// TIA Portal project "Inteligenta_szklarnia" (V15.1) (continued)
REGION Network 5
   RUNG wire#powerrail
      "Rolety"(Czy_automatyczny := wire#w1, Czy_manualny := wire#w2)
   END_RUNG
   RUNG wire#powerrail
      Contact( "HMI".Aktywacja_trybu_automatycznego )
   END_RUNG wire#w1
   RUNG wire#powerrail
      Contact( "HMI".Aktywacja_trybu_manualnego )
   END_RUNG wire#w2
   // the same network as SCL:
   "Rolety"(Czy_automatyczny := "HMI".Aktywacja_trybu_automatycznego,
            Czy_manualny := "HMI".Aktywacja_trybu_manualnego);
END_REGION

REGION Network 6
   RUNG wire#powerrail
      "Zapis_parametrow_trybu_auto"()
   END_RUNG
   // the same network as SCL:
   "Zapis_parametrow_trybu_auto"();
END_REGION

REGION Network 7
   RUNG wire#powerrail
      P_Contact(operand := "Clock_1Hz", bit := "marker_clock")
      "SYMULACJA"(counters := wire#w1)
   END_RUNG
   RUNG wire#powerrail
      I_Contact( "Clock_0.5Hz" )
   END_RUNG wire#w1
   // the same network as SCL:
   #_w1 := "Clock_1Hz" AND NOT "marker_clock";   // rising edge of "Clock_1Hz"
   "marker_clock" := "Clock_1Hz";
   IF #_w1 THEN "SYMULACJA"(counters := NOT "Clock_0.5Hz"); END_IF;
END_REGION

REGION Network 8
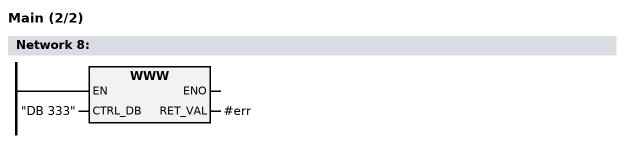
   #err := WWW(CTRL_DB := "DB 333");
END_REGION
END_ORGANIZATION_BLOCK

// folder: Archiwizacja_parametrow

FUNCTION "Archiwizacja_parametrow" : Void   // FC2, LAD
TITLE = Zapis parametrów oraz obliczanie z nich średniej każdego z ostatnich 7. dni
{ S7_Optimized_Access := 'TRUE' }
VERSION : 0.1
   VAR CONSTANT
      iterator : Int := 0;
   END_VAR
   VAR_TEMP   // added for the SCL form of the ladder/FBD networks
      _w1 : Bool;
   END_VAR
BEGIN

REGION Network 1: Zapis parametrów do bloku DB odbywa się co pół godziny. Po uruchomieniu sterownika pierwszy zapis nie odbywa się od razu, aby wykres nie przedstawiał parametrów, które nie były jeszcze regulowane. Odczytane wartości zapisywane są w tablicach w bloku DB.
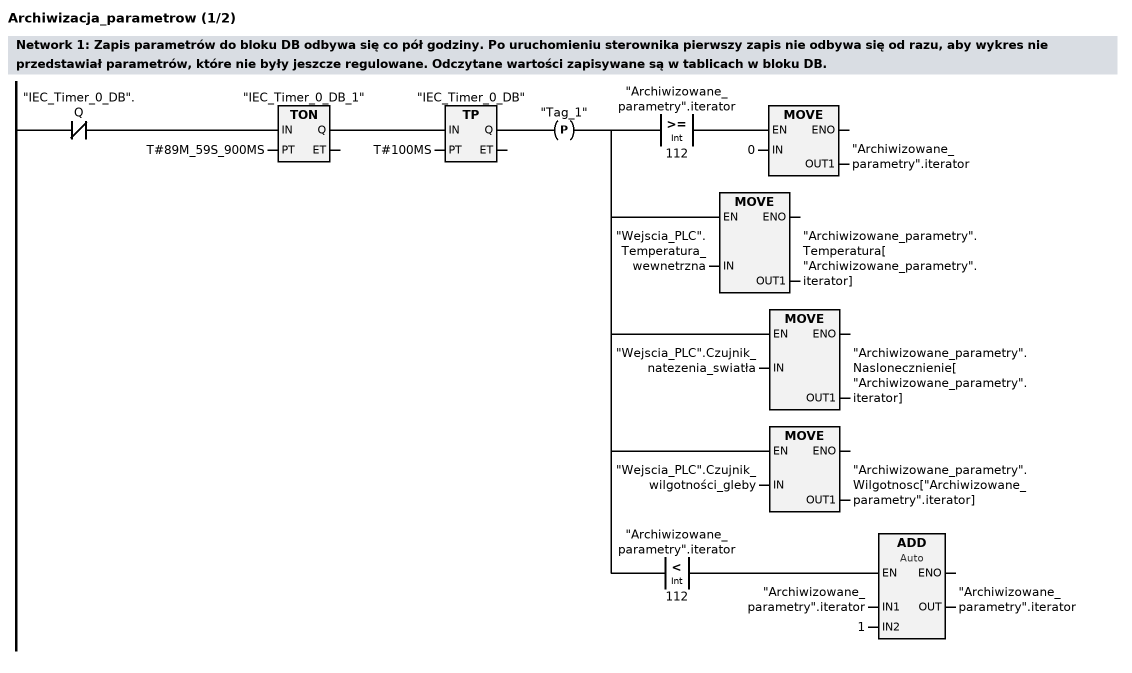
   "IEC_Timer_0_DB_1".TON(IN := NOT "IEC_Timer_0_DB".Q, PT := T#89M_59S_900MS);
   "IEC_Timer_0_DB".TP(IN := "IEC_Timer_0_DB_1".Q, PT := T#100MS);
   #_w1 := "IEC_Timer_0_DB".Q AND NOT "Tag_1";   // rising edge
   "Tag_1" := "IEC_Timer_0_DB".Q;
   IF #_w1 AND ("Archiwizowane_parametry".iterator >= 112) THEN
       "Archiwizowane_parametry".iterator := 0;
   END_IF;
   IF #_w1 THEN
       "Archiwizowane_parametry".Temperatura["Archiwizowane_parametry".iterator] := "Wejscia_PLC".Temperatura_wewnetrzna;
       "Archiwizowane_parametry".Naslonecznienie["Archiwizowane_parametry".iterator] := "Wejscia_PLC".Czujnik_natezenia_swiatła;
       "Archiwizowane_parametry".Wilgotnosc["Archiwizowane_parametry".iterator] := "Wejscia_PLC".Czujnik_wilgotności_gleby;
   END_IF;
   IF #_w1 AND ("Archiwizowane_parametry".iterator < 112) THEN
       "Archiwizowane_parametry".iterator := "Archiwizowane_parametry".iterator + 1;
   END_IF;
END_REGION

REGION Network 2: Zerowanie iteratora oraz zapisanych średnich w momencie zapisu kolejnych parametrów
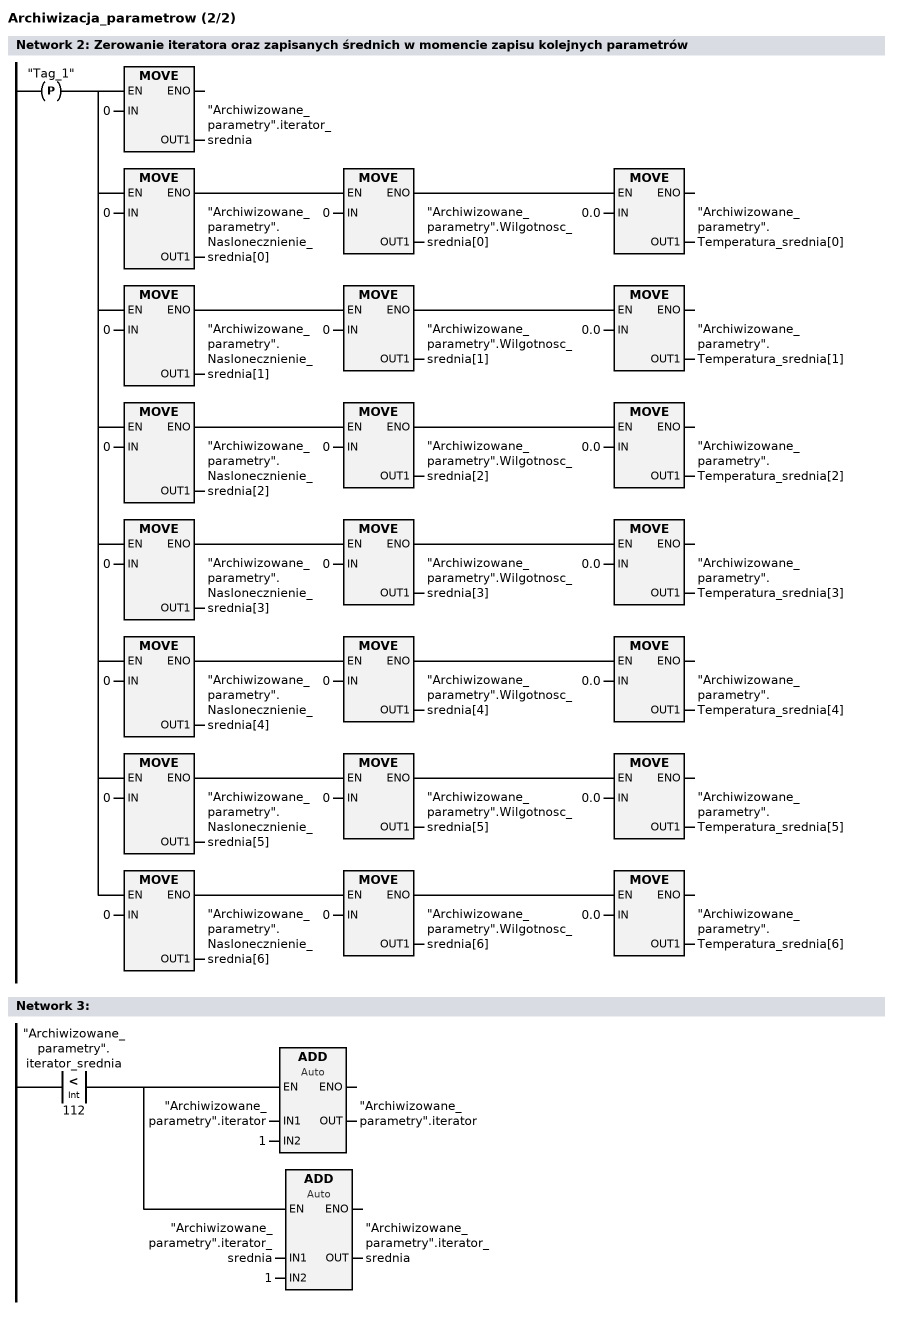
   RUNG wire#powerrail
      P_Trig( "Tag_1" )
      wire#w1
      { S7_GenerateENO := "TRUE" } Move(in := 0, out1 => "Archiwizowane_parametry".iterator_srednia)
   END_RUNG
   RUNG wire#w1
      { S7_GenerateENO := "TRUE" } Move(in := 0, out1 => "Archiwizowane_parametry".Naslonecznienie_srednia[0])
      { S7_GenerateENO := "TRUE" } Move(in := 0, out1 => "Archiwizowane_parametry".Wilgotnosc_srednia[0])
      { S7_GenerateENO := "TRUE" } Move(in := 0.0, out1 => "Archiwizowane_parametry".Temperatura_srednia[0])
   END_RUNG
   RUNG wire#w1
      { S7_GenerateENO := "TRUE" } Move(in := 0, out1 => "Archiwizowane_parametry".Naslonecznienie_srednia[1])
      { S7_GenerateENO := "TRUE" } Move(in := 0, out1 => "Archiwizowane_parametry".Wilgotnosc_srednia[1])
      { S7_GenerateENO := "TRUE" } Move(in := 0.0, out1 => "Archiwizowane_parametry".Temperatura_srednia[1])
   END_RUNG
   RUNG wire#w1
      { S7_GenerateENO := "TRUE" } Move(in := 0, out1 => "Archiwizowane_parametry".Naslonecznienie_srednia[2])
      { S7_GenerateENO := "TRUE" } Move(in := 0, out1 => "Archiwizowane_parametry".Wilgotnosc_srednia[2])
      { S7_GenerateENO := "TRUE" } Move(in := 0.0, out1 => "Archiwizowane_parametry".Temperatura_srednia[2])
   END_RUNG
   RUNG wire#w1
      { S7_GenerateENO := "TRUE" } Move(in := 0, out1 => "Archiwizowane_parametry".Naslonecznienie_srednia[3])
      { S7_GenerateENO := "TRUE" } Move(in := 0, out1 => "Archiwizowane_parametry".Wilgotnosc_srednia[3])
      { S7_GenerateENO := "TRUE" } Move(in := 0.0, out1 => "Archiwizowane_parametry".Temperatura_srednia[3])
   END_RUNG
   RUNG wire#w1
      { S7_GenerateENO := "TRUE" } Move(in := 0, out1 => "Archiwizowane_parametry".Naslonecznienie_srednia[4])
      { S7_GenerateENO := "TRUE" } Move(in := 0, out1 => "Archiwizowane_parametry".Wilgotnosc_srednia[4])
      { S7_GenerateENO := "TRUE" } Move(in := 0.0, out1 => "Archiwizowane_parametry".Temperatura_srednia[4])
   END_RUNG
   RUNG wire#w1
      { S7_GenerateENO := "TRUE" } Move(in := 0, out1 => "Archiwizowane_parametry".Naslonecznienie_srednia[5])
      { S7_GenerateENO := "TRUE" } Move(in := 0, out1 => "Archiwizowane_parametry".Wilgotnosc_srednia[5])
      { S7_GenerateENO := "TRUE" } Move(in := 0.0, out1 => "Archiwizowane_parametry".Temperatura_srednia[5])
   END_RUNG
   RUNG wire#w1
      { S7_GenerateENO := "TRUE" } Move(in := 0, out1 => "Archiwizowane_parametry".Naslonecznienie_srednia[6])
      { S7_GenerateENO := "TRUE" } Move(in := 0, out1 => "Archiwizowane_parametry".Wilgotnosc_srednia[6])
      { S7_GenerateENO := "TRUE" } Move(in := 0.0, out1 => "Archiwizowane_parametry".Temperatura_srednia[6])
   END_RUNG
   // the same network as SCL:
   // ENO of a box is taken as its EN; it also drops when the box reports an error
   #_w1 := NOT "Tag_1";   // rising edge
   "Tag_1" := TRUE;
   IF #_w1 THEN
       "Archiwizowane_parametry".iterator_srednia := 0;
       "Archiwizowane_parametry".Naslonecznienie_srednia[0] := 0;
       "Archiwizowane_parametry".Wilgotnosc_srednia[0] := 0;
       "Archiwizowane_parametry".Temperatura_srednia[0] := 0.0;
       "Archiwizowane_parametry".Naslonecznienie_srednia[1] := 0;
       "Archiwizowane_parametry".Wilgotnosc_srednia[1] := 0;
       "Archiwizowane_parametry".Temperatura_srednia[1] := 0.0;
       "Archiwizowane_parametry".Naslonecznienie_srednia[2] := 0;
       "Archiwizowane_parametry".Wilgotnosc_srednia[2] := 0;
       "Archiwizowane_parametry".Temperatura_srednia[2] := 0.0;
       "Archiwizowane_parametry".Naslonecznienie_srednia[3] := 0;
       "Archiwizowane_parametry".Wilgotnosc_srednia[3] := 0;
       "Archiwizowane_parametry".Temperatura_srednia[3] := 0.0;
       "Archiwizowane_parametry".Naslonecznienie_srednia[4] := 0;
       "Archiwizowane_parametry".Wilgotnosc_srednia[4] := 0;
       "Archiwizowane_parametry".Temperatura_srednia[4] := 0.0;
       "Archiwizowane_parametry".Naslonecznienie_srednia[5] := 0;
       "Archiwizowane_parametry".Wilgotnosc_srednia[5] := 0;
       "Archiwizowane_parametry".Temperatura_srednia[5] := 0.0;
       "Archiwizowane_parametry".Naslonecznienie_srednia[6] := 0;
       "Archiwizowane_parametry".Wilgotnosc_srednia[6] := 0;
       "Archiwizowane_parametry".Temperatura_srednia[6] := 0.0;
   END_IF;
END_REGION

REGION Network 3
   RUNG wire#powerrail
      { S7_Templates := "SrcType := Int" } LT_Contact(in1 := "Archiwizowane_parametry".iterator_srednia, in2 := 112)
      wire#w1
      { S7_GenerateENO := "TRUE" } Add(in1 := "Archiwizowane_parametry".iterator, in2 := 1, out => "Archiwizowane_parametry".iterator)
   END_RUNG
   RUNG wire#w1
      { S7_GenerateENO := "TRUE" } Add(in1 := "Archiwizowane_parametry".iterator_srednia, in2 := 1, out => "Archiwizowane_parametry".iterator_srednia)
   END_RUNG
   // the same network as SCL:
   IF "Archiwizowane_parametry".iterator_srednia < 112 THEN
       "Archiwizowane_parametry".iterator := "Archiwizowane_parametry".iterator + 1;
       "Archiwizowane_parametry".iterator_srednia := "Archiwizowane_parametry".iterator_srednia + 1;
   END_IF;
END_REGION
END_FUNCTION

// folder: LGF/4 Math operations

FUNCTION "LGF_RandomRange_Real" : Real   // FC10014, SCL
TITLE = LGF_RandomRange_Real
{ S7_Optimized_Access := 'TRUE' }
AUTHOR : Siemens_Digital_Industries
FAMILY : LGF
NAME : LGF_RandomRange_Real
// This function generates random numbers in defined limits (Datatype Real)
   VAR_INPUT
      minValue : Real;   // minimal Value random can reach / Minimum value of the range of the random number
      maxValue : Real;   // maximal Value random can reach / Maximum value of the range of the random number
   END_VAR
   VAR_OUTPUT
      error : Bool;   // Error if true
      status : Word;   // Status of the function
      subfunctionStatus : Word;   // Status or return value of called FB's, FCs and system blocks
   END_VAR
   VAR_TEMP
      tempTime : DTL;   // System time
      tempNanoSecondInDWord : DWord;   // UDINT converted to DWORD for access to individual bytes
      tempTimeStatus : Word;   // Status of the instruction RD_SYS_T
      tempRandomValue : DWord;   // Random-start-value
      tempNormReal : Real;   // normalized value
   END_VAR
   // Ret_Val : Returns random Real number in predefined range
   VAR CONSTANT
      ZERO : Real := 0.0;   // Zero value in case of error
      MAX_UDINT : UDInt := 4294967295;   // Maximum UDINT value
      SUB_STATUS_NO_ERROR : Word := 16#0000;   // Status: sub function call ends without error
      STATUS_FINISHED_NO_ERROR : Word := 16#0000;   // Status: Execution finished without errors
      ERR_MAX_LESS_MIN : Word := 16#8200;   // Error: The maximum limit number is smaller than the minimum limit number
      ERR_RD_SYS_T : Word := 16#8600;   // Error: System function Read system time returned an error
   END_VAR
BEGIN
   REGION Block info header
     //=============================================================================
     // SIEMENS AG / (c)Copyright 2017
     //-----------------------------------------------------------------------------
     // Title:            LGF_RandomRange_Real
     // Comment/Function: This function generates random numbers in defined limits (Datatype Real)
     // Library/Family:   LGF(Library General Functions)
     // Author:           Siemens Digital Industry Support
     // Tested with:      S7-PLCSIM Advanced V2.0 SP1
     // Engineering:      TIA Portal V15 Update 2
     // Restrictions:     ENO disabled - error handling done by error and status
     // Requirements:     PLC (S7-1200 / S7-1500)
     //-------------------------------------------------------------------------------
     // Change log table:
     // Version  | Date       | Expert in charge       | Changes applied
     //----------|------------|------------------------|------------------------------
     // 01.00.00 19.08.2015  Siemens Industry Online Support
     //                      First released version
     // 01.00.01 02.01.2017  Siemens Industry Online Support
     //                      Upgrade: TIA Portal V14 Update 1
     // 01.00.02 02.03.2017  Siemens Industry Online Support
     //                      Bugfix: FC number
     // 01.00.03 17.08.2018  Siemens Industry Online Support
     //                      Upgrade: TIA V15 Update 2
     // 01.00.04 23.11.2018  Siemens Industry Online Support
     //                      Upgrade: TIA V15.1
     // 01.01.00 13.11.2019  Siemens Industry Presales Support
     //                      Renamed from "LGF_RandomReal" to "LGF_RandomRange_Real"
     //                      Regions, commens and costants are added
     // 03.00.00 23.04.2020  Siemens Industry Support
     //                      Set version to V3.0.0, harmonize the version of the whole library
     //=============================================================================
   END_REGION

   REGION Validation
     // Check if the maximal Value is less than the minimal value
     IF (#minValue > #maxValue) THEN
       #error := true;
       #status := #ERR_MAX_LESS_MIN;
       #subfunctionStatus := #SUB_STATUS_NO_ERROR;
       #LGF_RandomRange_Real := #ZERO;
       RETURN;
     END_IF;

     // Read system time
     #tempTimeStatus := INT_TO_WORD(RD_SYS_T(#tempTime));

     // Check return variable for error
     IF (#tempTimeStatus <> #SUB_STATUS_NO_ERROR) THEN
       #error := true;
       #status := #ERR_RD_SYS_T;
       #subfunctionStatus := #tempTimeStatus;
       #LGF_RandomRange_Real := #ZERO;
       RETURN;
     END_IF;
   END_REGION

   REGION Calculating random number
     // Converting to double word so individual bytes can be addressed
     #tempNanoSecondInDWord := UDINT_TO_DWORD(#tempTime.NANOSECOND);

     // Calculate a random-start-value depending on the time
     #tempRandomValue.%B3 := #tempNanoSecondInDWord.%B0;
     #tempRandomValue.%B2 := #tempNanoSecondInDWord.%B1;
     #tempRandomValue.%B1 := #tempNanoSecondInDWord.%B2;
     #tempRandomValue.%B0 := #tempNanoSecondInDWord.%B3;

     // Norm the calculated random number: 0.0 <= #tempNormReal <= 1.0
     #tempNormReal := UDINT_TO_REAL(DWORD_TO_UDINT(#tempRandomValue)) / UDINT_TO_REAL(#MAX_UDINT);

     // Scale the tempNormReal to be in the range of maxValue and minValue
     #LGF_RandomRange_Real := ((#tempNormReal * (#maxValue - #minValue) + (#minValue)));

     #error := false;
     #status := #STATUS_FINISHED_NO_ERROR;
     #subfunctionStatus := #SUB_STATUS_NO_ERROR;
     // ENO mechanism is not used
     ENO := TRUE;
   END_REGION
END_FUNCTION

// ===== PLC "PLC_do_symulacji"  CPU 1214C AC/DC/Rly =====

VAR_GLOBAL   // PLC tag table "Default tag table"
   "Tag_1" AT %M0.0 : Bool;
   "System_Byte" AT %MB1 : Byte;
   "FirstScan" AT %M1.0 : Bool;
   "DiagStatusUpdate" AT %M1.1 : Bool;
   "AlwaysTRUE" AT %M1.2 : Bool;
   "AlwaysFALSE" AT %M1.3 : Bool;
   "Tag_2" AT %M0.1 : Bool;
   "Clock_Byte" AT %MB30 : Byte;
   "Clock_10Hz" AT %M30.0 : Bool;
   "Clock_5Hz" AT %M30.1 : Bool;
   "Clock_2.5Hz" AT %M30.2 : Bool;
   "Clock_2Hz" AT %M30.3 : Bool;
   "Clock_1.25Hz" AT %M30.4 : Bool;
   "Clock_1Hz" AT %M30.5 : Bool;
   "Clock_0.625Hz" AT %M30.6 : Bool;
   "Clock_0.5Hz" AT %M30.7 : Bool;
   "marker_clock" AT %M0.2 : Bool;
   "marker_counter" AT %M0.3 : Bool;
   "wartosc_rolet_sym" AT %MW2 : Int;
   "swiatlo_bez_rolet" AT %MW4 : Int;
   "Alarm_active" AT %M6.0 : Bool;
   "Tag_3" AT %M0.4 : Bool;
END_VAR

VAR_GLOBAL   // PLC tag table "wyjscia"
   "Grzałka" AT %Q0.0 : Bool;
   "Wentylator" AT %Q0.1 : Bool;
   "Pompa_zraszacze" AT %Q0.2 : Bool;   // Pompa zraszaczy, które odpowiadają za wilgotność powietrza w szklarni
   "Rolety_zamykanie" AT %Q0.4 : Bool;
   "Alarm_ostrzegwaczy" AT %Q0.5 : Bool;
   "Siłownik_okien_otwieranie" AT %Q0.6 : Bool;
   "Siłownik_okien_zamykanie" AT %Q0.7 : Bool;
   "Rolety_otwieranie" AT %Q0.3 : Bool;
   "Pompa_podlewanie" AT %Q1.0 : Bool;   // Pompa podlewania kropelkowego, która odpowiada za wilgotność gleby
END_VAR

DATA_BLOCK "Wejscia_PLC"   // DB1
{ S7_Optimized_Access := 'TRUE' }
VERSION : 0.1
   VAR
      Czujnik_wilgotności_powietrza : Int;   // Czujnik wilgotności powietrza w szklarni
      Czujnik_wilgotności_gleby : Int;   // Czujnik wilgotności gleby w szklarni
      Temperatura_wewnetrzna : Real;   // Temperatura wewnątrz szklarni
      Czujnik_natezenia_swiatła : Int;   // Czujnik natężenia światła wewnątrz szklarni
      Czujnik_wiatru : Int;   // Czujnik prędkości wiatru poza szklarnią
      Wewnetrzny_czujnik_CO2 : Int;   // Czujnik stężenia dwutlenku węgla w szklarni
      Stopien_zasloniecia_rolet : Int;   // Stopień zasłonięcia rolet w szklarni (przyjęty przedział 0-100%)
      Temperatura_zewnetrzna : Real;   // Temperatura mierzona na zewnątrz, poza szklarnią. Typ Int, ponieważ nie jest wymagana taka dokładność jak w pomiarze temperatury wewnętrznej.
      Zewnetrzny_czujnik_CO2 : Int;   // Czujnik stężenia dwutlenku węgla poza szklarnią
      czujnik_wilgotnosci_zewnetrzny : Int := 50;   // Potrzebny w ramach symulacji realnych warunkow
   END_VAR
BEGIN
END_DATA_BLOCK

DATA_BLOCK "HMI"   // DB2
{ S7_Optimized_Access := 'TRUE' }
VERSION : 0.1
   VAR
      nazwa_receptury : String;
      System_okien_auto : Bool;   // Wł/wył system okien w trybie automatycznym
      Przycisk_zraszacze_manual : Bool;   // Przycisk pompy zraszaczy w trybie manualnym
      Przycisk_podlewanie_manual : Bool;   // Przycisk pompy podlewania w trybie manualnym
      Przycisk_grzanie_manual : Bool;   // Przycisk grzałki w trybie manualnym
      Przycisk_wentylacja_manual : Bool;   // Przycisk wentylacji w trybie manualnym
      Otwarcie_okien_manual : Bool;   // Ustawiony w trybie manualnym otwarcie okien
      Stopien_zasloniecia_rolet_manual : Int;   // Ustawiony w trybie manualnym stopień zasłonięcia rolet
      Temperatura_auto : Real := 22.0;   // Nastawiona temeratura w trybie automatycznym
      Naslonecznienie_auto : Int := 1000;   // Nastawiona wartość nasłonecznienia w trybie automatycznym
      Wilgotnosc_powietrza_auto : Int := 50;   // Nastawiona wartość wilgotności powietrza w trybie automatycznym
      Poziom_CO2_auto : Int := 800;   // Nastawiona wartość stężenia CO2 w trybie automatycznym
      Wilgotnosc_gleby_auto : Int := 60;   // Nastawiona wartość wilgotności gleby w trybie automatycznym
      Przycisk_zatwierdz_auto : Bool;   // Przycisk zatwierdzający wcześniej wybrane ustawienia trybu automatycznego
      Przycisk_zatwierdz_zapis_receptury : Bool;   // Przycisk zatwierdzający wcześniej wybrane ustawienia trybu zapisania receptury
      Przycisk_zatwierdz_wybor_receptury : Bool;   // Przycisk zatwierdzający wcześniej wybrane ustawienia trybu receptury
      Numer_ekranu_HMI : Int;   // Numer aktualnie otwartego ekranu w HMI
      Aktywacja_trybu_manualnego : Bool;
      Aktywacja_trybu_automatycznego : Bool;
      Aktywacja_trybu_Receptur : Bool;
      Aktywacja_trybu_zapis_Receptur : Bool;
      Reset_Trybow : Bool;
   END_VAR
BEGIN
END_DATA_BLOCK

DATA_BLOCK "Tryb_auto_parametry"   // DB7
{ S7_Optimized_Access := 'TRUE' }
VERSION : 0.1
   VAR
      Temperatura : Real;
      Naslonecznienie : Int;
      Wilgotnosc_powietrza : Int;
      Wilgotnosc_gleby : Int;
      System_okien : Bool;
      Stezenie_co2 : Int;
   END_VAR
BEGIN
END_DATA_BLOCK

DATA_BLOCK "Alarmy"   // DB9
{ S7_Optimized_Access := 'TRUE' }
VERSION : 0.1
   VAR
      alarmW : Word;
      Warning_niska_temp_1 : Bool;
      Warning_wysoka_temp_1 : Bool;
      Warning_nieprawidlowe_CO2_1 : Bool;
   END_VAR
BEGIN
END_DATA_BLOCK

// folder: Archiwizacja_parametrow

DATA_BLOCK "Archiwizowane_parametry"   // DB4
{ S7_Optimized_Access := 'TRUE' }
VERSION : 0.1
   VAR
      Temperatura : Array[0..111] of Real;
      Wilgotnosc : Array[0..111] of Int;
      Naslonecznienie : Array[0..111] of Int;
      iterator : Int := 0;   // Iterator służący do zapisu danych w odpowiednich komórkach tablicy.
      Temperatura_srednia : Array[0..6] of Real;
      Wilgotnosc_srednia : Array[0..6] of Int;
      Naslonecznienie_srednia : Array[0..6] of Int;
      iterator_srednia : Int := 0;   // Iterator służący do zapisu danych w odpowiednich komórkach tablicy.
      dzielnik : Int;   // Ilość zsumowanych parametrów w średniej
      Temperatura_suma : Array[0..6] of Real;
      Wilgotnosc_suma : Array[0..6] of Int;
      Naslonecznienie_suma : Array[0..6] of Int;
   END_VAR
BEGIN
   Naslonecznienie[0] := -1;
   Naslonecznienie[1] := -1;
   Temperatura[0] := -20.0;
   Temperatura[1] := -20.0;
   Temperatura[2] := -20.0;
   Temperatura[3] := -20.0;
   Temperatura[4] := -20.0;
   Temperatura[5] := -20.0;
   Temperatura[12] := -20.0;
   Temperatura[13] := -20.0;
   Temperatura[14] := -20.0;
   Temperatura[15] := -20.0;
   Temperatura[16] := -20.0;
   Temperatura[17] := -20.0;
   Temperatura[6] := -20.0;
   Temperatura[7] := -20.0;
   Temperatura[8] := -20.0;
   Temperatura[9] := -20.0;
   Temperatura[10] := -20.0;
   Temperatura[11] := -20.0;
   Temperatura[18] := -20.0;
   Temperatura[19] := -20.0;
   Temperatura[20] := -20.0;
   Temperatura[21] := -20.0;
   Temperatura[22] := -20.0;
   Temperatura[23] := -20.0;
   Temperatura[24] := -20.0;
   Temperatura[25] := -20.0;
   Temperatura[26] := -20.0;
   Temperatura[27] := -20.0;
   Temperatura[28] := -20.0;
   Temperatura[29] := -20.0;
   Temperatura[30] := -20.0;
   Temperatura[31] := -20.0;
   Temperatura[32] := -20.0;
   Temperatura[33] := -20.0;
   Temperatura[34] := -20.0;
   Temperatura[35] := -20.0;
   Temperatura[36] := -20.0;
   Temperatura[37] := -20.0;
   Temperatura[38] := -20.0;
   Temperatura[39] := -20.0;
   Temperatura[40] := -20.0;
   Temperatura[41] := -20.0;
   Temperatura[42] := -20.0;
   Temperatura[43] := -20.0;
   Temperatura[44] := -20.0;
   Temperatura[45] := -20.0;
   Temperatura[46] := -20.0;
   Temperatura[47] := -20.0;
   Temperatura[48] := -20.0;
   Temperatura[49] := -20.0;
   Temperatura[50] := -20.0;
   Temperatura[51] := -20.0;
   Temperatura[52] := -20.0;
   Temperatura[53] := -20.0;
   Temperatura[54] := -20.0;
   Temperatura[55] := -20.0;
   Temperatura[56] := -20.0;
   Temperatura[57] := -20.0;
   Temperatura[58] := -20.0;
   Temperatura[59] := -20.0;
   Temperatura[60] := -20.0;
   Temperatura[61] := -20.0;
   Temperatura[62] := -20.0;
   Temperatura[63] := -20.0;
   Temperatura[64] := -20.0;
   Temperatura[65] := -20.0;
   Temperatura[66] := -20.0;
   Temperatura[67] := -20.0;
   Temperatura[68] := -20.0;
   Temperatura[69] := -20.0;
   Temperatura[70] := -20.0;
   Temperatura[71] := -20.0;
   Temperatura[72] := -20.0;
   Temperatura[73] := -20.0;
   Temperatura[74] := -20.0;
   Temperatura[75] := -20.0;
   Temperatura[76] := -20.0;
   Temperatura[77] := -20.0;
   Temperatura[78] := -20.0;
   Temperatura[79] := -20.0;
   Temperatura[80] := -20.0;
   Temperatura[81] := -20.0;
   Temperatura[82] := -20.0;
   Temperatura[83] := -20.0;
   Temperatura[84] := -20.0;
   Temperatura[85] := -20.0;
   Temperatura[86] := -20.0;
   Temperatura[87] := -20.0;
   Temperatura[88] := -20.0;
   Temperatura[89] := -20.0;
   Temperatura[90] := -20.0;
   Temperatura[91] := -20.0;
   Temperatura[92] := -20.0;
   Temperatura[93] := -20.0;
   Temperatura[94] := -20.0;
   Temperatura[95] := -20.0;
   Temperatura[96] := -20.0;
   Temperatura[97] := -20.0;
   Temperatura[98] := -20.0;
   Temperatura[99] := -20.0;
   Temperatura[100] := -20.0;
   Temperatura[101] := -20.0;
   Temperatura[102] := -20.0;
   Temperatura[103] := -20.0;
   Temperatura[104] := -20.0;
   Temperatura[105] := -20.0;
   Temperatura[106] := -20.0;
   Temperatura[107] := -20.0;
   Temperatura[108] := -20.0;
   Temperatura[109] := -20.0;
   Temperatura[110] := -20.0;
   Temperatura[111] := -20.0;
   Wilgotnosc[0] := -1;
   Wilgotnosc[1] := -1;
   Wilgotnosc[2] := -1;
   Wilgotnosc[3] := -1;
   Wilgotnosc[4] := -1;
   Wilgotnosc[5] := -1;
   Wilgotnosc[6] := -1;
   Wilgotnosc[7] := -1;
   Wilgotnosc[8] := -1;
   Wilgotnosc[9] := -1;
   Wilgotnosc[10] := -1;
   Wilgotnosc[11] := -1;
   Wilgotnosc[12] := -1;
   Wilgotnosc[13] := -1;
   Wilgotnosc[14] := -1;
   Wilgotnosc[15] := -1;
   Wilgotnosc[16] := -1;
   Wilgotnosc[17] := -1;
   Wilgotnosc[18] := -1;
   Wilgotnosc[19] := -1;
   Wilgotnosc[20] := -1;
   Wilgotnosc[21] := -1;
   Wilgotnosc[22] := -1;
   Wilgotnosc[23] := -1;
   Wilgotnosc[24] := -1;
   Wilgotnosc[25] := -1;
   Wilgotnosc[26] := -1;
   Wilgotnosc[27] := -1;
   Wilgotnosc[28] := -1;
   Wilgotnosc[29] := -1;
   Wilgotnosc[30] := -1;
   Wilgotnosc[31] := -1;
   Wilgotnosc[32] := -1;
   Wilgotnosc[33] := -1;
   Wilgotnosc[34] := -1;
   Wilgotnosc[35] := -1;
   Wilgotnosc[36] := -1;
   Wilgotnosc[37] := -1;
   Wilgotnosc[38] := -1;
   Wilgotnosc[39] := -1;
   Wilgotnosc[40] := -1;
   Wilgotnosc[41] := -1;
   Wilgotnosc[42] := -1;
   Wilgotnosc[43] := -1;
   Wilgotnosc[44] := -1;
   Wilgotnosc[45] := -1;
   Wilgotnosc[46] := -1;
   Wilgotnosc[47] := -1;
   Wilgotnosc[48] := -1;
   Wilgotnosc[49] := -1;
   Wilgotnosc[50] := -1;
   Wilgotnosc[51] := -1;
   Wilgotnosc[52] := -1;
   Wilgotnosc[53] := -1;
   Wilgotnosc[54] := -1;
   Wilgotnosc[55] := -1;
   Wilgotnosc[56] := -1;
   Wilgotnosc[57] := -1;
   Wilgotnosc[58] := -1;
   Wilgotnosc[59] := -1;
   Wilgotnosc[60] := -1;
   Wilgotnosc[61] := -1;
   Wilgotnosc[62] := -1;
   Wilgotnosc[63] := -1;
   Wilgotnosc[64] := -1;
   Wilgotnosc[65] := -1;
   Wilgotnosc[66] := -1;
   Wilgotnosc[67] := -1;
   Wilgotnosc[68] := -1;
   Wilgotnosc[69] := -1;
   Wilgotnosc[70] := -1;
   Wilgotnosc[71] := -1;
   Wilgotnosc[72] := -1;
   Wilgotnosc[73] := -1;
   Wilgotnosc[74] := -1;
   Wilgotnosc[75] := -1;
   Wilgotnosc[76] := -1;
   Wilgotnosc[77] := -1;
   Wilgotnosc[78] := -1;
   Wilgotnosc[79] := -1;
   Wilgotnosc[80] := -1;
   Wilgotnosc[81] := -1;
   Wilgotnosc[82] := -1;
   Wilgotnosc[83] := -1;
   Wilgotnosc[84] := -1;
   Wilgotnosc[85] := -1;
   Wilgotnosc[86] := -1;
   Wilgotnosc[87] := -1;
   Wilgotnosc[88] := -1;
   Wilgotnosc[89] := -1;
   Wilgotnosc[90] := -1;
   Wilgotnosc[91] := -1;
   Wilgotnosc[92] := -1;
   Wilgotnosc[93] := -1;
   Wilgotnosc[94] := -1;
   Wilgotnosc[95] := -1;
   Wilgotnosc[96] := -1;
   Wilgotnosc[97] := -1;
   Wilgotnosc[98] := -1;
   Wilgotnosc[99] := -1;
   Wilgotnosc[100] := -1;
   Wilgotnosc[101] := -1;
   Wilgotnosc[102] := -1;
   Wilgotnosc[103] := -1;
   Wilgotnosc[104] := -1;
   Wilgotnosc[105] := -1;
   Wilgotnosc[106] := -1;
   Wilgotnosc[107] := -1;
   Wilgotnosc[108] := -1;
   Wilgotnosc[109] := -1;
   Wilgotnosc[110] := -1;
   Wilgotnosc[111] := -1;
   Naslonecznienie[2] := -1;
   Naslonecznienie[3] := -1;
   Naslonecznienie[4] := -1;
   Naslonecznienie[5] := -1;
   Naslonecznienie[6] := -1;
   Naslonecznienie[7] := -1;
   Naslonecznienie[8] := -1;
   Naslonecznienie[9] := -1;
   Naslonecznienie[10] := -1;
   Naslonecznienie[11] := -1;
   Naslonecznienie[12] := -1;
   Naslonecznienie[13] := -1;
   Naslonecznienie[14] := -1;
   Naslonecznienie[15] := -1;
   Naslonecznienie[16] := -1;
   Naslonecznienie[17] := -1;
   Naslonecznienie[18] := -1;
   Naslonecznienie[19] := -1;
   Naslonecznienie[20] := -1;
   Naslonecznienie[21] := -1;
   Naslonecznienie[22] := -1;
   Naslonecznienie[23] := -1;
   Naslonecznienie[24] := -1;
   Naslonecznienie[25] := -1;
   Naslonecznienie[26] := -1;
   Naslonecznienie[27] := -1;
   Naslonecznienie[28] := -1;
   Naslonecznienie[29] := -1;
   Naslonecznienie[30] := -1;
   Naslonecznienie[31] := -1;
   Naslonecznienie[32] := -1;
   Naslonecznienie[33] := -1;
   Naslonecznienie[34] := -1;
   Naslonecznienie[35] := -1;
   Naslonecznienie[36] := -1;
   Naslonecznienie[37] := -1;
   Naslonecznienie[38] := -1;
   Naslonecznienie[39] := -1;
   Naslonecznienie[40] := -1;
   Naslonecznienie[41] := -1;
   Naslonecznienie[42] := -1;
   Naslonecznienie[43] := -1;
   Naslonecznienie[44] := -1;
   Naslonecznienie[45] := -1;
   Naslonecznienie[46] := -1;
   Naslonecznienie[47] := -1;
   Naslonecznienie[48] := -1;
   Naslonecznienie[49] := -1;
   Naslonecznienie[50] := -1;
   Naslonecznienie[51] := -1;
   Naslonecznienie[52] := -1;
   Naslonecznienie[53] := -1;
   Naslonecznienie[54] := -1;
   Naslonecznienie[55] := -1;
   Naslonecznienie[56] := -1;
   Naslonecznienie[57] := -1;
   Naslonecznienie[58] := -1;
   Naslonecznienie[59] := -1;
   Naslonecznienie[60] := -1;
   Naslonecznienie[61] := -1;
   Naslonecznienie[62] := -1;
   Naslonecznienie[63] := -1;
   Naslonecznienie[64] := -1;
   Naslonecznienie[65] := -1;
   Naslonecznienie[66] := -1;
   Naslonecznienie[67] := -1;
   Naslonecznienie[68] := -1;
   Naslonecznienie[69] := -1;
   Naslonecznienie[70] := -1;
   Naslonecznienie[71] := -1;
   Naslonecznienie[72] := -1;
   Naslonecznienie[73] := -1;
   Naslonecznienie[74] := -1;
   Naslonecznienie[75] := -1;
   Naslonecznienie[76] := -1;
   Naslonecznienie[77] := -1;
   Naslonecznienie[78] := -1;
   Naslonecznienie[79] := -1;
   Naslonecznienie[80] := -1;
   Naslonecznienie[81] := -1;
   Naslonecznienie[82] := -1;
   Naslonecznienie[83] := -1;
   Naslonecznienie[84] := -1;
   Naslonecznienie[85] := -1;
   Naslonecznienie[86] := -1;
   Naslonecznienie[87] := -1;
   Naslonecznienie[88] := -1;
   Naslonecznienie[89] := -1;
   Naslonecznienie[90] := -1;
   Naslonecznienie[91] := -1;
   Naslonecznienie[92] := -1;
   Naslonecznienie[93] := -1;
   Naslonecznienie[94] := -1;
   Naslonecznienie[95] := -1;
   Naslonecznienie[96] := -1;
   Naslonecznienie[97] := -1;
   Naslonecznienie[98] := -1;
   Naslonecznienie[99] := -1;
   Naslonecznienie[100] := -1;
   Naslonecznienie[101] := -1;
   Naslonecznienie[102] := -1;
   Naslonecznienie[103] := -1;
   Naslonecznienie[104] := -1;
   Naslonecznienie[105] := -1;
   Naslonecznienie[106] := -1;
   Naslonecznienie[107] := -1;
   Naslonecznienie[108] := -1;
   Naslonecznienie[109] := -1;
   Naslonecznienie[110] := -1;
   Naslonecznienie[111] := -1;
   // Temperatura_srednia[0] : Dzień 1.
END_DATA_BLOCK

// folder: System blocks/Program resources

DATA_BLOCK "IEC_Counter_0_DB_1"   // DB3
{ S7_Optimized_Access := 'TRUE' }
AUTHOR : Simatic
FAMILY : IEC
NAME : CNTR
VERSION : 1.0
// stored: InstanceOfName IEC_COUNTER
"IEC_COUNTER"
BEGIN
END_DATA_BLOCK

DATA_BLOCK "IEC_Timer_0_DB"   // DB5
{ S7_Optimized_Access := 'TRUE' }
AUTHOR : Simatic
FAMILY : IEC
NAME : IEC_TMR
VERSION : 1.0
// stored: InstanceOfName IEC_TIMER
"IEC_TIMER"
BEGIN
END_DATA_BLOCK

DATA_BLOCK "IEC_Timer_0_DB_1"   // DB6
{ S7_Optimized_Access := 'TRUE' }
AUTHOR : Simatic
FAMILY : IEC
NAME : IEC_TMR
VERSION : 1.0
// stored: InstanceOfName IEC_TIMER
"IEC_TIMER"
BEGIN
END_DATA_BLOCK

DATA_BLOCK "IEC_Timer_0_DB_2"   // DB8
{ S7_Optimized_Access := 'TRUE' }
AUTHOR : Simatic
FAMILY : IEC
NAME : IEC_TMR
VERSION : 1.0
// stored: InstanceOfName IEC_TIMER
"IEC_TIMER"
BEGIN
END_DATA_BLOCK

DATA_BLOCK "IEC_Timer_0_DB_5"   // DB10
{ S7_Optimized_Access := 'TRUE' }
AUTHOR : Simatic
FAMILY : IEC
NAME : IEC_TMR
VERSION : 1.0
// stored: InstanceOfName IEC_TIMER
"IEC_TIMER"
BEGIN
END_DATA_BLOCK

DATA_BLOCK "IEC_Timer_0_DB_3"   // DB11
{ S7_Optimized_Access := 'TRUE' }
AUTHOR : Simatic
FAMILY : IEC
NAME : IEC_TMR
VERSION : 1.0
// stored: InstanceOfName IEC_TIMER
"IEC_TIMER"
BEGIN
END_DATA_BLOCK

DATA_BLOCK "IEC_Counter_0_DB"   // DB12
{ S7_Optimized_Access := 'TRUE' }
AUTHOR : Simatic
FAMILY : IEC
NAME : CNTR
VERSION : 1.0
// stored: InstanceOfName IEC_COUNTER
"IEC_COUNTER"
BEGIN
END_DATA_BLOCK

DATA_BLOCK "IEC_Counter_0_DB_2"   // DB13
{ S7_Optimized_Access := 'TRUE' }
AUTHOR : Simatic
FAMILY : IEC
NAME : CNTR
VERSION : 1.0
// stored: InstanceOfName IEC_COUNTER
"IEC_COUNTER"
BEGIN
END_DATA_BLOCK

// folder: (top level)

FUNCTION "Rolety" : Void   // FC1, LAD
{ S7_Optimized_Access := 'TRUE' }
VERSION : 0.1
   VAR_INPUT
      Czy_automatyczny : Bool;
      Czy_manualny : Bool;
   END_VAR
BEGIN

REGION Network 1: Warunki otwierania rolet w trybie automatycznym i manualnym
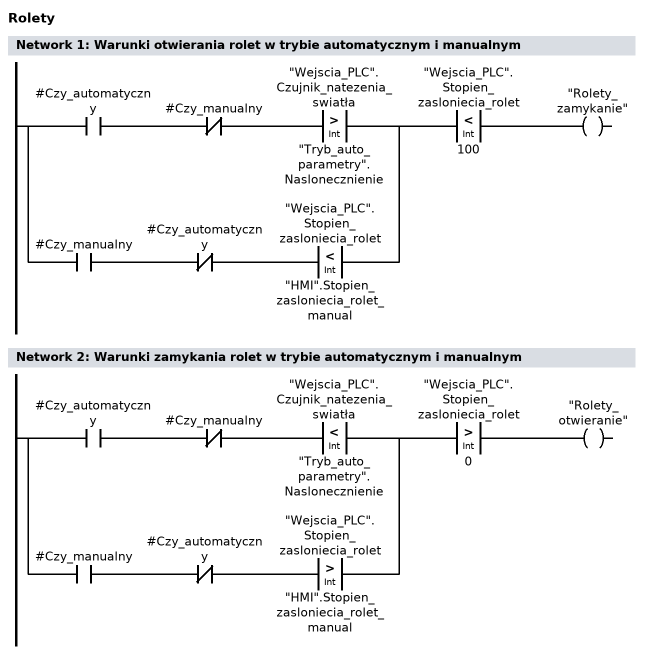
   RUNG wire#powerrail
      Contact( #Czy_automatyczny )
      I_Contact( #Czy_manualny )
      { S7_Templates := "SrcType := Int" } GT_Contact(in1 := "Wejscia_PLC".Czujnik_natezenia_swiatła, in2 := "Tryb_auto_parametry".Naslonecznienie)
      wire#w1
      { S7_Templates := "SrcType := Int" } LT_Contact(in1 := "Wejscia_PLC".Stopien_zasloniecia_rolet, in2 := 100)
      Coil( "Rolety_zamykanie" )
   END_RUNG
   RUNG wire#powerrail
      Contact( #Czy_manualny )
      I_Contact( #Czy_automatyczny )
      { S7_Templates := "SrcType := Int" } LT_Contact(in1 := "Wejscia_PLC".Stopien_zasloniecia_rolet, in2 := "HMI".Stopien_zasloniecia_rolet_manual)
   END_RUNG wire#w1
   // the same network as SCL:
   "Rolety_zamykanie" := ((#Czy_automatyczny AND NOT #Czy_manualny AND ("Wejscia_PLC".Czujnik_natezenia_swiatła > "Tryb_auto_parametry".Naslonecznienie)) OR (#Czy_manualny AND NOT #Czy_automatyczny AND ("Wejscia_PLC".Stopien_zasloniecia_rolet < "HMI".Stopien_zasloniecia_rolet_manual))) AND ("Wejscia_PLC".Stopien_zasloniecia_rolet < 100);
END_REGION

REGION Network 2: Warunki zamykania rolet w trybie automatycznym i manualnym
   RUNG wire#powerrail
      Contact( #Czy_automatyczny )
      I_Contact( #Czy_manualny )
      { S7_Templates := "SrcType := Int" } LT_Contact(in1 := "Wejscia_PLC".Czujnik_natezenia_swiatła, in2 := "Tryb_auto_parametry".Naslonecznienie)
      wire#w1
      { S7_Templates := "SrcType := Int" } GT_Contact(in1 := "Wejscia_PLC".Stopien_zasloniecia_rolet, in2 := 0)
      Coil( "Rolety_otwieranie" )
   END_RUNG
   RUNG wire#powerrail
      Contact( #Czy_manualny )
      I_Contact( #Czy_automatyczny )
      { S7_Templates := "SrcType := Int" } GT_Contact(in1 := "Wejscia_PLC".Stopien_zasloniecia_rolet, in2 := "HMI".Stopien_zasloniecia_rolet_manual)
   END_RUNG wire#w1
   // the same network as SCL:
   "Rolety_otwieranie" := ((#Czy_automatyczny AND NOT #Czy_manualny AND ("Wejscia_PLC".Czujnik_natezenia_swiatła < "Tryb_auto_parametry".Naslonecznienie)) OR (#Czy_manualny AND NOT #Czy_automatyczny AND ("Wejscia_PLC".Stopien_zasloniecia_rolet > "HMI".Stopien_zasloniecia_rolet_manual))) AND ("Wejscia_PLC".Stopien_zasloniecia_rolet > 0);
END_REGION
END_FUNCTION

FUNCTION "Sterowanie_grzalka_wentylator" : Void   // FC3, LAD
{ S7_Optimized_Access := 'TRUE' }
VERSION : 0.1
   VAR_INPUT
      czy_manualny : Bool;
      czy_automatyczny : Bool;
   END_VAR
   VAR_TEMP
      Histereza_minus : Real;   // Wartość zadanej temperatury zmieniona o dolną wartość hiterezy
      Histereza_plus : Real;   // Wartość zadanej temperatury zmieniona o górną wartość hiterezy
   END_VAR
   VAR CONSTANT
      Wartosc_histerezy : Real := 1.0;
   END_VAR
   VAR_TEMP   // added for the SCL form of the ladder/FBD networks
      _w1 : Bool;
   END_VAR
BEGIN

REGION Network 1: Sterowanie wentylatorem w trybie automatycznym i manualnym
   // Gdy uruchomiony jest tryb automatyczny, wartość temperatury w szklarni powinna się mieścić w zakresie temperatury nastawionej +- wartość histerezy. Gdy jest ona za wysoka uruchamiany jest wentylator. W trybie manualnym włączany jest on od razu po naciśnięciu przycisku do niego przypisanego.
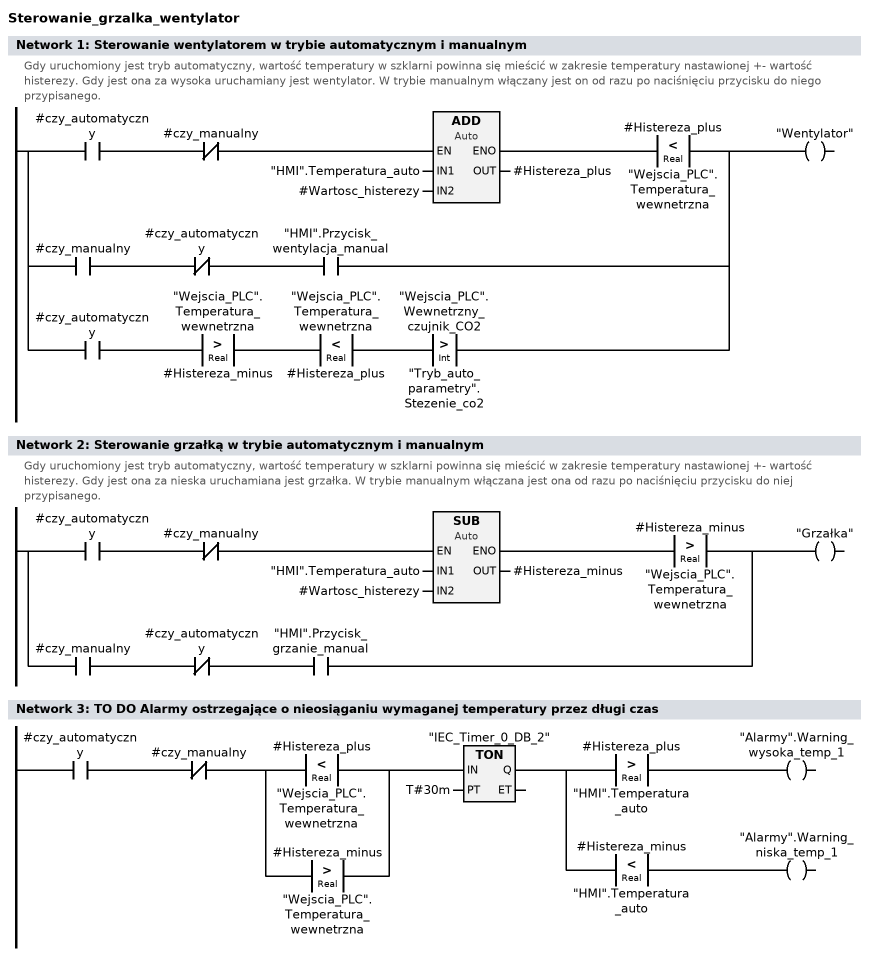
   RUNG wire#powerrail
      Contact( #czy_automatyczny )
      I_Contact( #czy_manualny )
      Add(in1 := "HMI".Temperatura_auto, in2 := #Wartosc_histerezy, out => #Histereza_plus)
      { S7_Templates := "SrcType := Real" } LT_Contact(in1 := #Histereza_plus, in2 := "Wejscia_PLC".Temperatura_wewnetrzna)
      wire#w1
      Coil( "Wentylator" )
   END_RUNG
   RUNG wire#powerrail
      Contact( #czy_manualny )
      I_Contact( #czy_automatyczny )
      Contact( "HMI".Przycisk_wentylacja_manual )
   END_RUNG wire#w1
   RUNG wire#powerrail
      Contact( #czy_automatyczny )
      { S7_Templates := "SrcType := Real" } GT_Contact(in1 := "Wejscia_PLC".Temperatura_wewnetrzna, in2 := #Histereza_minus)
      { S7_Templates := "SrcType := Real" } LT_Contact(in1 := "Wejscia_PLC".Temperatura_wewnetrzna, in2 := #Histereza_plus)
      { S7_Templates := "SrcType := Int" } GT_Contact(in1 := "Wejscia_PLC".Wewnetrzny_czujnik_CO2, in2 := "Tryb_auto_parametry".Stezenie_co2)
   END_RUNG wire#w1
   // the same network as SCL:
   #_w1 := #czy_automatyczny AND NOT #czy_manualny;
   IF #_w1 THEN #Histereza_plus := "HMI".Temperatura_auto + #Wartosc_histerezy; END_IF;
   "Wentylator" := (#_w1 AND (#Histereza_plus < "Wejscia_PLC".Temperatura_wewnetrzna)) OR (#czy_manualny AND NOT #czy_automatyczny AND "HMI".Przycisk_wentylacja_manual) OR (#czy_automatyczny AND ("Wejscia_PLC".Temperatura_wewnetrzna > #Histereza_minus) AND ("Wejscia_PLC".Temperatura_wewnetrzna < #Histereza_plus) AND ("Wejscia_PLC".Wewnetrzny_czujnik_CO2 > "Tryb_auto_parametry".Stezenie_co2));
END_REGION

REGION Network 2: Sterowanie grzałką w trybie automatycznym i manualnym
   // Gdy uruchomiony jest tryb automatyczny, wartość temperatury w szklarni powinna się mieścić w zakresie temperatury nastawionej +- wartość histerezy. Gdy jest ona za nieska uruchamiana jest grzałka. W trybie manualnym włączana jest ona od razu po naciśnięciu przycisku do niej przypisanego.
   RUNG wire#powerrail
      Contact( #czy_automatyczny )
      I_Contact( #czy_manualny )
      Sub(in1 := "HMI".Temperatura_auto, in2 := #Wartosc_histerezy, out => #Histereza_minus)
      { S7_Templates := "SrcType := Real" } GT_Contact(in1 := #Histereza_minus, in2 := "Wejscia_PLC".Temperatura_wewnetrzna)
      wire#w1
      Coil( "Grzałka" )
   END_RUNG
   RUNG wire#powerrail
      Contact( #czy_manualny )
      I_Contact( #czy_automatyczny )
      Contact( "HMI".Przycisk_grzanie_manual )
   END_RUNG wire#w1
   // the same network as SCL:
   #_w1 := #czy_automatyczny AND NOT #czy_manualny;
   IF #_w1 THEN #Histereza_minus := "HMI".Temperatura_auto - #Wartosc_histerezy; END_IF;
   "Grzałka" := (#_w1 AND (#Histereza_minus > "Wejscia_PLC".Temperatura_wewnetrzna)) OR (#czy_manualny AND NOT #czy_automatyczny AND "HMI".Przycisk_grzanie_manual);
END_REGION

REGION Network 3: TO DO Alarmy ostrzegające o nieosiąganiu wymaganej temperatury przez długi czas
   "IEC_Timer_0_DB_2".TON(IN := #czy_automatyczny AND NOT #czy_manualny AND ((#Histereza_plus < "Wejscia_PLC".Temperatura_wewnetrzna) OR (#Histereza_minus > "Wejscia_PLC".Temperatura_wewnetrzna)),
                          PT := T#30m);
   "Alarmy".Warning_wysoka_temp_1 := "IEC_Timer_0_DB_2".Q AND (#Histereza_plus > "HMI".Temperatura_auto);
   "Alarmy".Warning_niska_temp_1 := "IEC_Timer_0_DB_2".Q AND (#Histereza_minus < "HMI".Temperatura_auto);
END_REGION
END_FUNCTION

FUNCTION "Zapis_parametrow_trybu_auto" : Void   // FC4, LAD
{ S7_Optimized_Access := 'TRUE' }
VERSION : 0.1
BEGIN

REGION Network 1: Zapis wybranych na HMI parametrów, aby zostały one stałe do kolejnego zatwierdzenia ich zmiany.
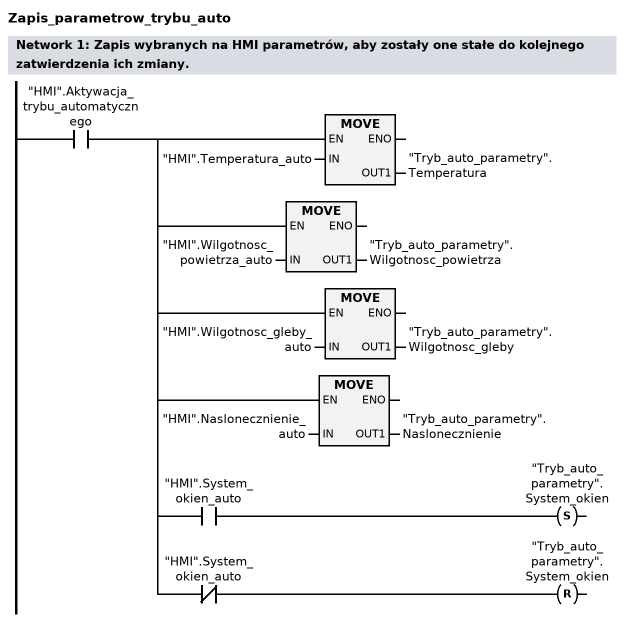
   RUNG wire#powerrail
      Contact( "HMI".Aktywacja_trybu_automatycznego )
      wire#w1
      Move(in := "HMI".Temperatura_auto, out1 => "Tryb_auto_parametry".Temperatura)
   END_RUNG
   RUNG wire#w1
      Move(in := "HMI".Wilgotnosc_powietrza_auto, out1 => "Tryb_auto_parametry".Wilgotnosc_powietrza)
   END_RUNG
   RUNG wire#w1
      Move(in := "HMI".Wilgotnosc_gleby_auto, out1 => "Tryb_auto_parametry".Wilgotnosc_gleby)
   END_RUNG
   RUNG wire#w1
      Move(in := "HMI".Naslonecznienie_auto, out1 => "Tryb_auto_parametry".Naslonecznienie)
   END_RUNG
   RUNG wire#w1
      Contact( "HMI".System_okien_auto )
      S_Coil( "Tryb_auto_parametry".System_okien )
   END_RUNG
   RUNG wire#w1
      I_Contact( "HMI".System_okien_auto )
      R_Coil( "Tryb_auto_parametry".System_okien )
   END_RUNG
   // the same network as SCL:
   IF "HMI".Aktywacja_trybu_automatycznego THEN
       "Tryb_auto_parametry".Temperatura := "HMI".Temperatura_auto;
       "Tryb_auto_parametry".Wilgotnosc_powietrza := "HMI".Wilgotnosc_powietrza_auto;
       "Tryb_auto_parametry".Wilgotnosc_gleby := "HMI".Wilgotnosc_gleby_auto;
       "Tryb_auto_parametry".Naslonecznienie := "HMI".Naslonecznienie_auto;
   END_IF;
   IF "HMI".Aktywacja_trybu_automatycznego AND "HMI".System_okien_auto THEN
       "Tryb_auto_parametry".System_okien := TRUE;
   END_IF;
   IF "HMI".Aktywacja_trybu_automatycznego AND NOT "HMI".System_okien_auto THEN
       "Tryb_auto_parametry".System_okien := FALSE;
   END_IF;
END_REGION
END_FUNCTION

FUNCTION "Jaki_Tryb" : Void   // FC5, LAD
{ S7_Optimized_Access := 'TRUE' }
VERSION : 0.1
BEGIN

REGION Network 1: Reset trybu auto jesli wykryje jakikolwiek inny tryb
